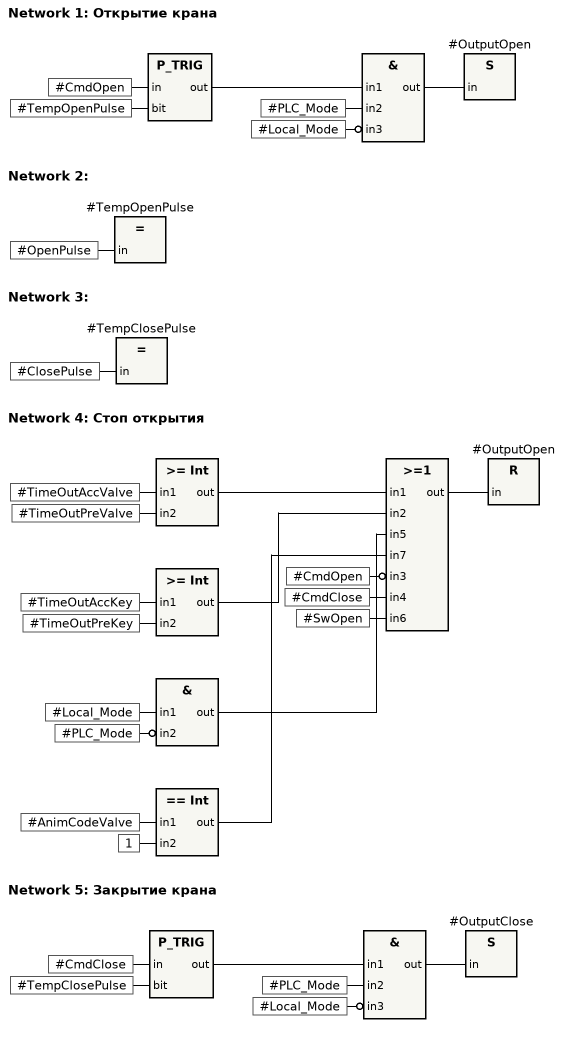
   #_w1 := #CmdOpen AND NOT #TempOpenPulse;   // rising edge
   #TempOpenPulse := #CmdOpen;
   IF #_w1 AND #PLC_Mode AND NOT #Local_Mode THEN #OutputOpen := TRUE; END_IF;
END_REGION

REGION Network 2
   #TempOpenPulse := #OpenPulse;
END_REGION

REGION Network 3
   #TempClosePulse := #ClosePulse;
END_REGION

REGION Network 4: Стоп открытия
   IF (#TimeOutAccValve >= #TimeOutPreValve) OR (#TimeOutAccKey >= #TimeOutPreKey) OR (#Local_Mode AND NOT #PLC_Mode) OR (#AnimCodeValve = 1) OR NOT #CmdOpen OR #CmdClose OR #SwOpen THEN
       #OutputOpen := FALSE;
   END_IF;
END_REGION

REGION Network 5: Закрытие крана
   #_w1 := #CmdClose AND NOT #TempClosePulse;   // rising edge
   #TempClosePulse := #CmdClose;
   IF #_w1 AND #PLC_Mode AND NOT #Local_Mode THEN #OutputClose := TRUE; END_IF;
END_REGION

REGION Network 6: Стоп закрытия
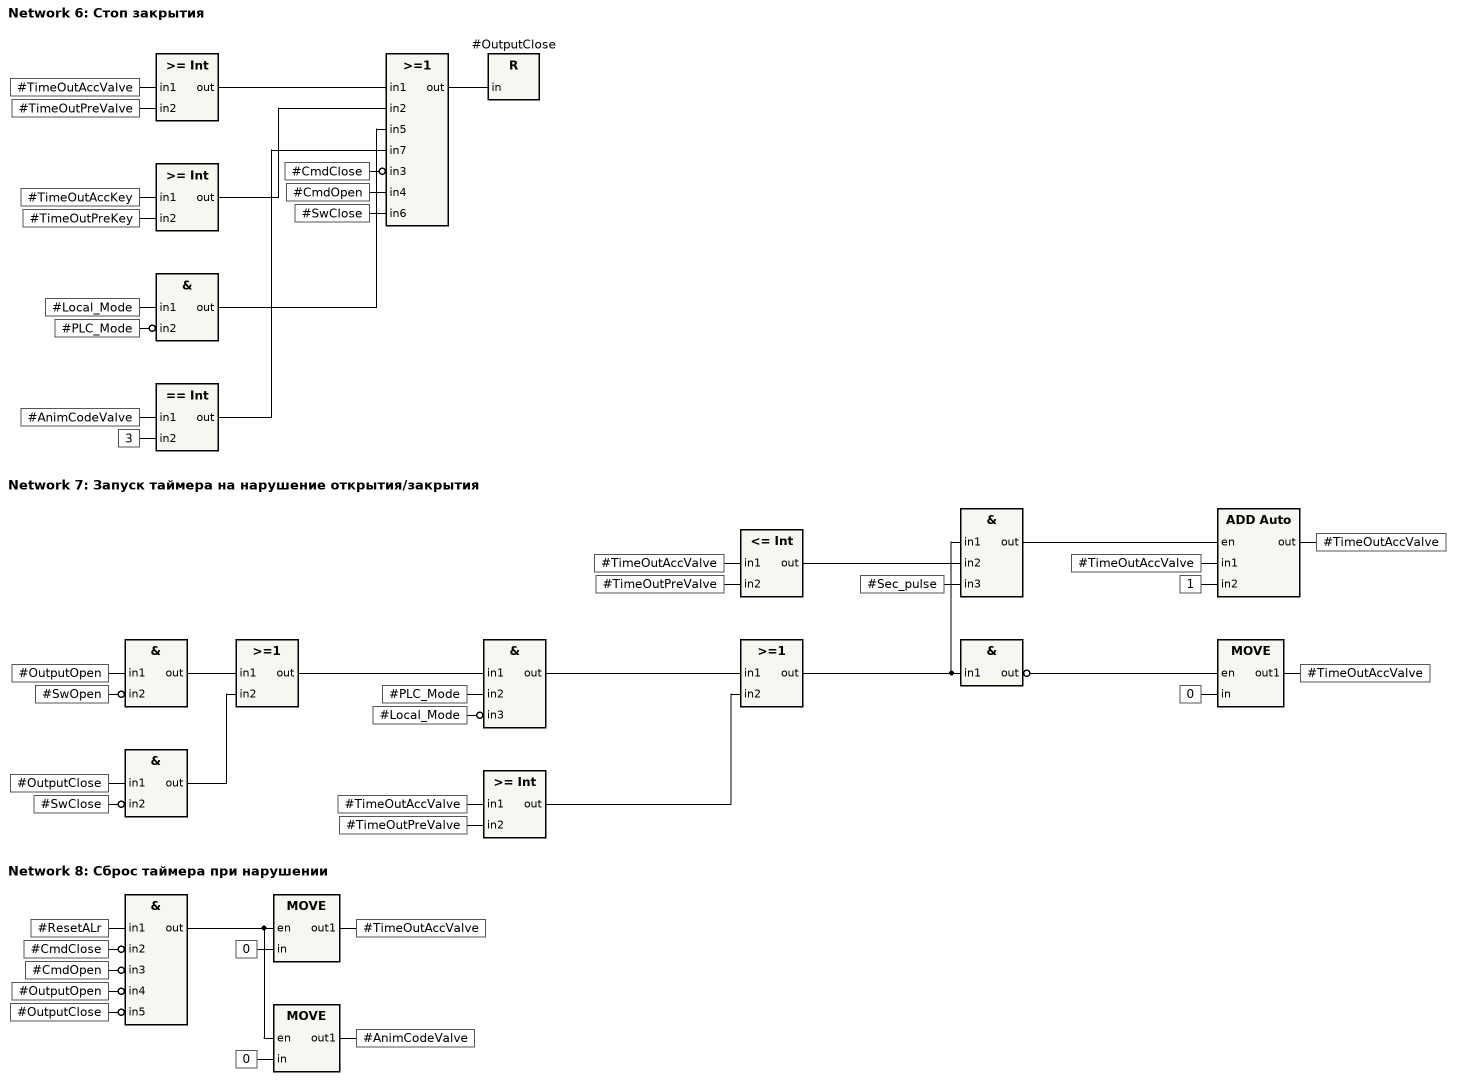
   IF (#TimeOutAccValve >= #TimeOutPreValve) OR (#TimeOutAccKey >= #TimeOutPreKey) OR (#Local_Mode AND NOT #PLC_Mode) OR (#AnimCodeValve = 3) OR NOT #CmdClose OR #CmdOpen OR #SwClose THEN
       #OutputClose := FALSE;
   END_IF;
END_REGION

REGION Network 7: Запуск таймера на нарушение открытия/закрытия
   #_w1 := (((#OutputOpen AND NOT #SwOpen) OR (#OutputClose AND NOT #SwClose)) AND #PLC_Mode AND NOT #Local_Mode) OR (#TimeOutAccValve >= #TimeOutPreValve);
   IF #_w1 AND (#TimeOutAccValve <= #TimeOutPreValve) AND #Sec_pulse THEN
       #TimeOutAccValve := #TimeOutAccValve + 1;
   END_IF;
   IF NOT #_w1 THEN #TimeOutAccValve := 0; END_IF;
END_REGION

REGION Network 8: Сброс таймера при нарушении
   IF #ResetALr AND NOT #CmdClose AND NOT #CmdOpen AND NOT #OutputOpen AND NOT #OutputClose THEN
       #TimeOutAccValve := 0;
       #AnimCodeValve := 0;
   END_IF;
END_REGION

REGION Network 9: Код анимации состояния крана
   // 0-Нейтральное
   // 1-Открыт
   // 2-Открывается
   // 3-Закрыт
   // 4-Закрывается
   // 10- Нарушения открытия
   // 11- Нарушения закрытия
   // 12- Открытие без команды
   // 13- Закрытие без команды
   // 14- Оба датчика включены
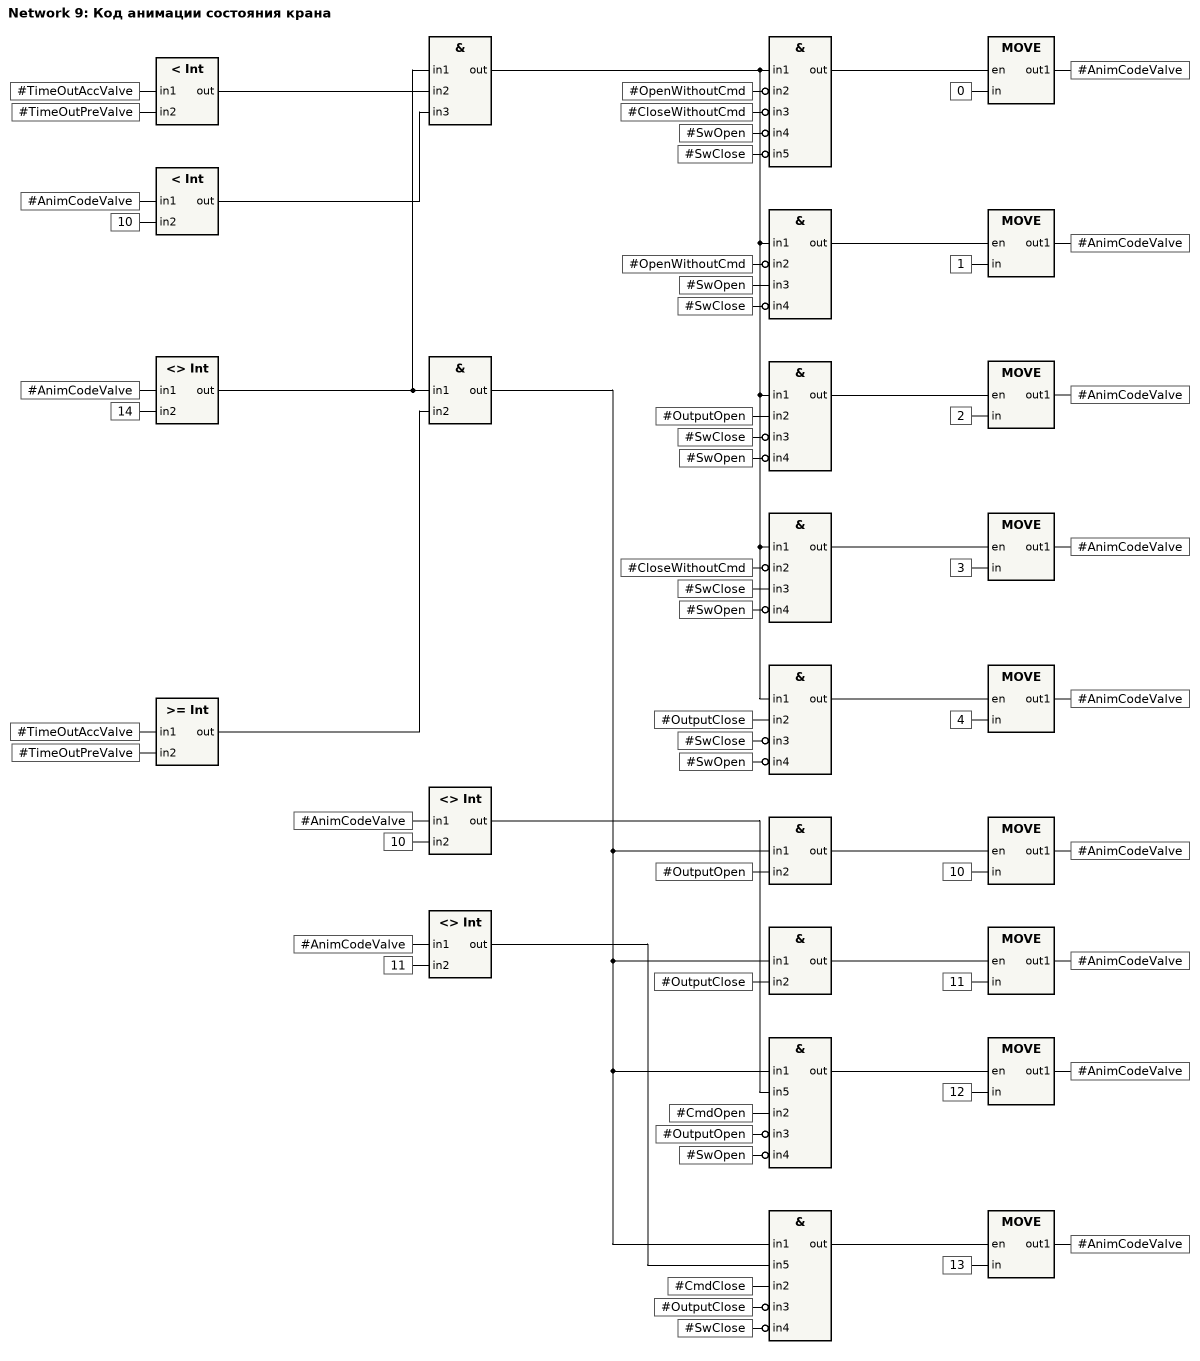
   #_w1 := #AnimCodeValve <> 14;
   #_w2 := #_w1 AND (#TimeOutAccValve < #TimeOutPreValve) AND (#AnimCodeValve < 10);
   IF #_w2 AND NOT #OpenWithoutCmd AND NOT #CloseWithoutCmd AND NOT #SwOpen AND NOT #SwClose THEN
       #AnimCodeValve := 0;
   END_IF;
   IF #_w2 AND NOT #OpenWithoutCmd AND #SwOpen AND NOT #SwClose THEN #AnimCodeValve := 1; END_IF;
   IF #_w2 AND #OutputOpen AND NOT #SwClose AND NOT #SwOpen THEN #AnimCodeValve := 2; END_IF;
   IF #_w2 AND NOT #CloseWithoutCmd AND #SwClose AND NOT #SwOpen THEN #AnimCodeValve := 3; END_IF;
   IF #_w2 AND #OutputClose AND NOT #SwClose AND NOT #SwOpen THEN #AnimCodeValve := 4; END_IF;
   #_w3 := #_w1 AND (#TimeOutAccValve >= #TimeOutPreValve);
   IF #_w3 AND #OutputOpen THEN #AnimCodeValve := 10; END_IF;
   IF #_w3 AND #OutputClose THEN #AnimCodeValve := 11; END_IF;
   IF #_w3 AND (#AnimCodeValve <> 10) AND #CmdOpen AND NOT #OutputOpen AND NOT #SwOpen THEN
       #AnimCodeValve := 12;
   END_IF;
   IF #_w3 AND (#AnimCodeValve <> 11) AND #CmdClose AND NOT #OutputClose AND NOT #SwClose THEN
       #AnimCodeValve := 13;
   END_IF;
END_REGION

REGION Network 10: Два датчика включены
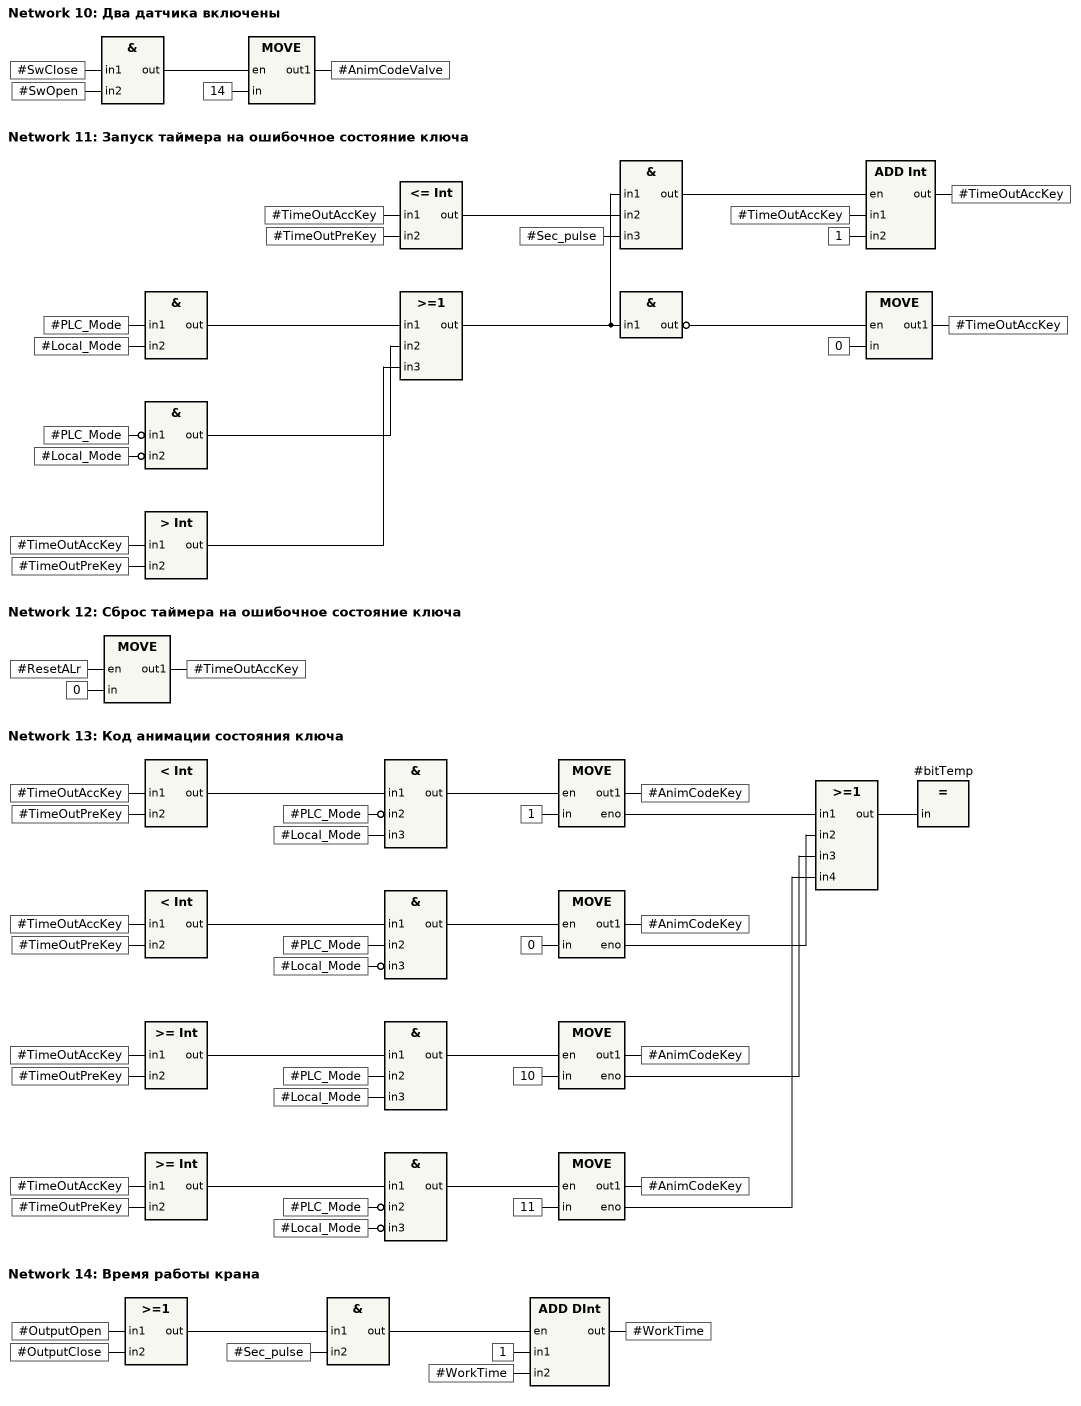
   IF #SwClose AND #SwOpen THEN #AnimCodeValve := 14; END_IF;
END_REGION

REGION Network 11: Запуск таймера на ошибочное состояние ключа
   #_w1 := (#PLC_Mode AND #Local_Mode) OR (NOT #PLC_Mode AND NOT #Local_Mode) OR (#TimeOutAccKey > #TimeOutPreKey);
   IF #_w1 AND (#TimeOutAccKey <= #TimeOutPreKey) AND #Sec_pulse THEN
       #TimeOutAccKey := #TimeOutAccKey + 1;
   END_IF;
   IF NOT #_w1 THEN #TimeOutAccKey := 0; END_IF;
END_REGION

REGION Network 12: Сброс таймера на ошибочное состояние ключа
   IF #ResetALr THEN #TimeOutAccKey := 0; END_IF;
END_REGION

REGION Network 13: Код анимации состояния ключа
   // ENO of a box is taken as its EN; it also drops when the box reports an error
   #_w1 := (#TimeOutAccKey < #TimeOutPreKey) AND NOT #PLC_Mode AND #Local_Mode;
   IF #_w1 THEN #AnimCodeKey := 1; END_IF;
   #_w2 := (#TimeOutAccKey < #TimeOutPreKey) AND #PLC_Mode AND NOT #Local_Mode;
   IF #_w2 THEN #AnimCodeKey := 0; END_IF;
   #_w3 := (#TimeOutAccKey >= #TimeOutPreKey) AND #PLC_Mode AND #Local_Mode;
   IF #_w3 THEN #AnimCodeKey := 10; END_IF;
   #_w4 := (#TimeOutAccKey >= #TimeOutPreKey) AND NOT #PLC_Mode AND NOT #Local_Mode;
   IF #_w4 THEN #AnimCodeKey := 11; END_IF;
   #bitTemp := #_w1 OR #_w2 OR #_w3 OR #_w4;
END_REGION

REGION Network 14: Время работы крана
   IF (#OutputOpen OR #OutputClose) AND #Sec_pulse THEN #WorkTime := 1 + #WorkTime; END_IF;
END_REGION

REGION Network 15: Сброс времени работы мотора
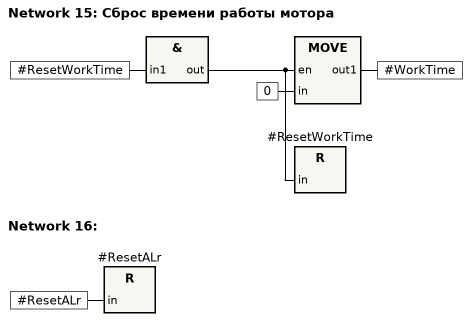
   IF #ResetWorkTime THEN
       #WorkTime := 0;
       #ResetWorkTime := FALSE;
   END_IF;
END_REGION

REGION Network 16
   IF #ResetALr THEN #ResetALr := FALSE; END_IF;
END_REGION
END_FUNCTION

FUNCTION "106_Analog_Type" : Void   // FC106, FBD
{ S7_Optimized_Access := 'TRUE' }
VERSION : 0.1
   VAR_INPUT
      Input : Int;
      Eng_Hi : Real;
      Eng_Lo : Real;
      Sp_HiHi : Real;
      Sp_Hi : Real;
      Sp_Lo : Real;
      Sp_LoLo : Real;
   END_VAR
   VAR_OUTPUT
      Value : Real;
      Alm_HiHi : Bool;
      Alm_Hi : Bool;
      Alm_Lo : Bool;
      Alm_LoLo : Bool;
      AnimCode : Int;
      OpenLoop : Bool;
      ShortCircuit : Bool;
   END_VAR
   VAR_TEMP
      Val_Conv : Real;
      Val_Temp : Real;
      Bool_Tmp : Bool;
      Input_Tmp : Int;
      tAlm_HiHi : Bool;
      tAlm_Hi : Bool;
      tAlm_Lo : Bool;
      tAlm_LoLo : Bool;
      tOpenLoop : Bool;
      tShortCircuit : Bool;
   END_VAR
BEGIN

REGION Network 1
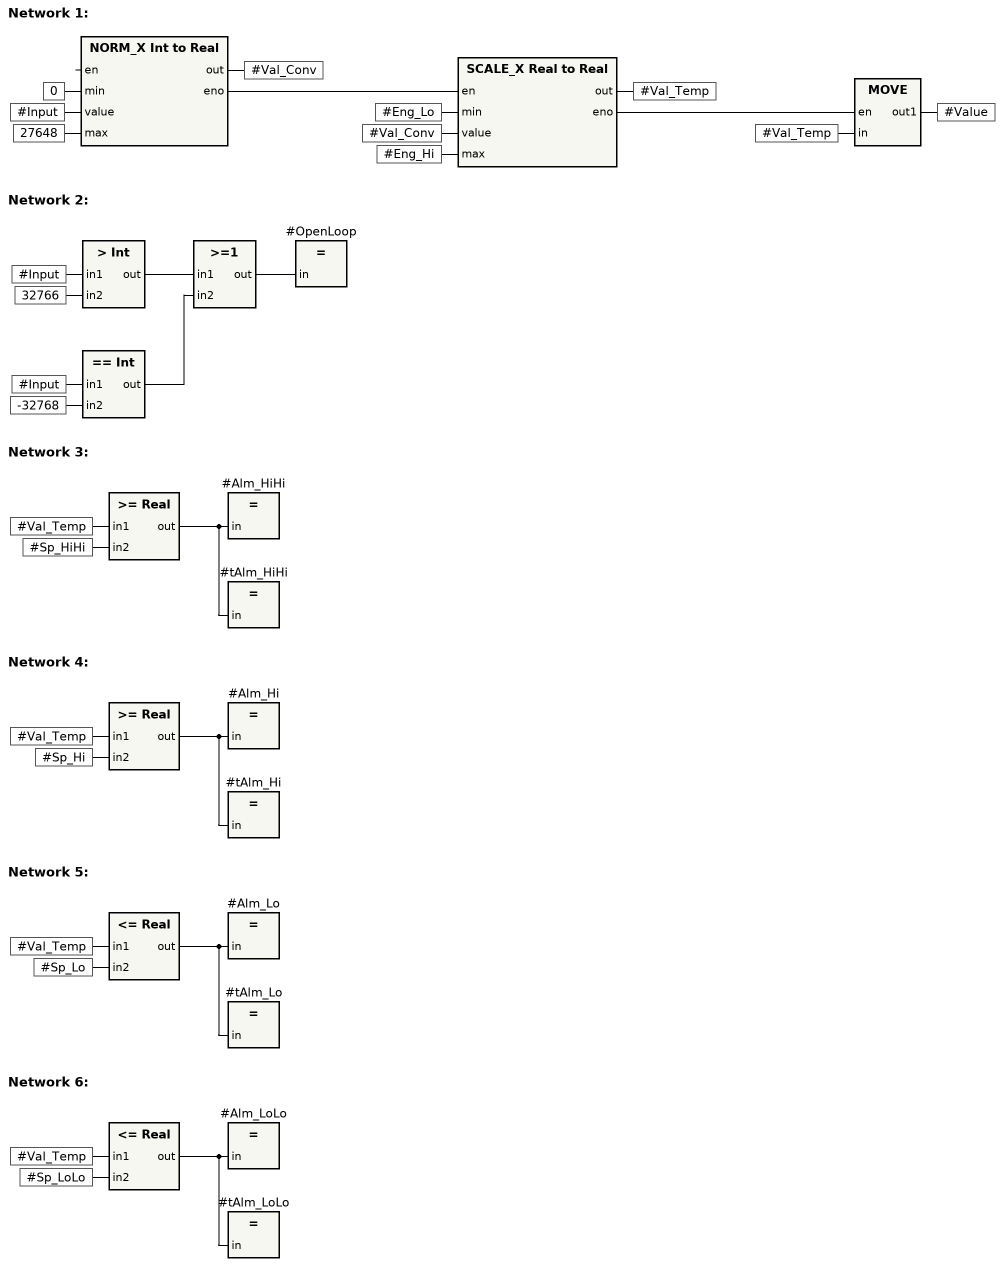
   // ENO of a box is taken as its EN; it also drops when the box reports an error
   #Val_Conv := NORM_X(MIN := 0, VALUE := #Input, MAX := 27648);
   #Val_Temp := SCALE_X(MIN := #Eng_Lo, VALUE := #Val_Conv, MAX := #Eng_Hi);
   #Value := #Val_Temp;
END_REGION

REGION Network 2
   #OpenLoop := (#Input > 32766) OR (#Input = (-32768));
END_REGION

REGION Network 3
   #Alm_HiHi := #Val_Temp >= #Sp_HiHi;
   #tAlm_HiHi := #Alm_HiHi;
END_REGION

REGION Network 4
   #Alm_Hi := #Val_Temp >= #Sp_Hi;
   #tAlm_Hi := #Alm_Hi;
END_REGION

REGION Network 5
   #Alm_Lo := #Val_Temp <= #Sp_Lo;
   #tAlm_Lo := #Alm_Lo;
END_REGION

REGION Network 6
   #Alm_LoLo := #Val_Temp <= #Sp_LoLo;
   #tAlm_LoLo := #Alm_LoLo;
END_REGION

REGION Network 7
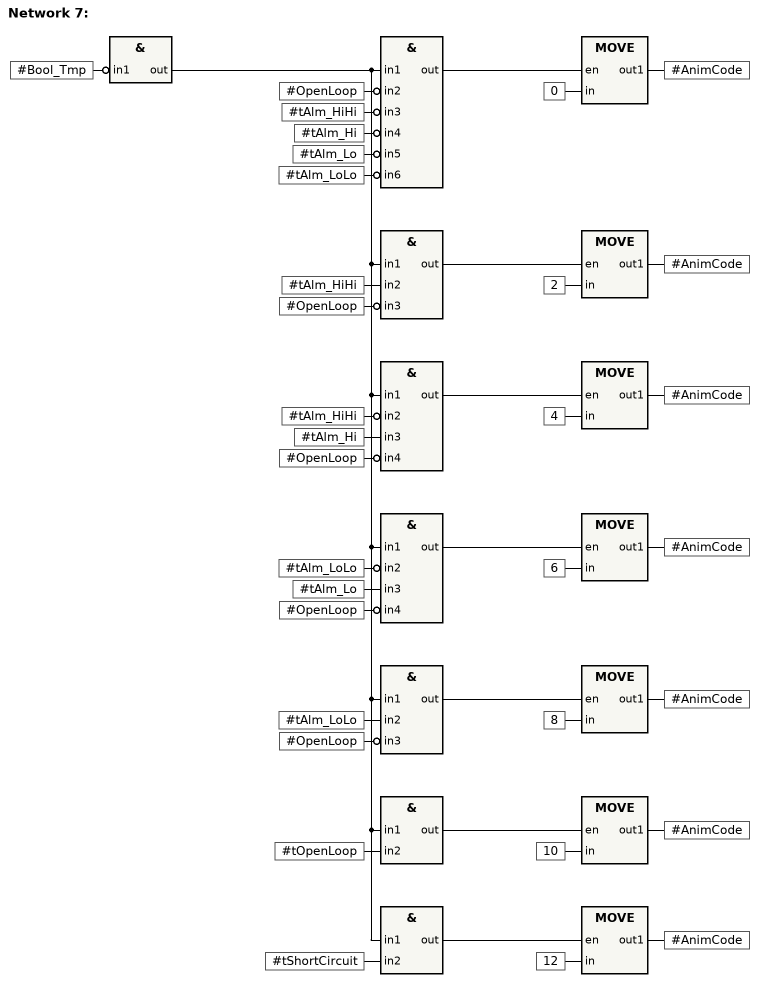
   IF NOT #Bool_Tmp AND NOT #OpenLoop AND NOT #tAlm_HiHi AND NOT #tAlm_Hi AND NOT #tAlm_Lo AND NOT #tAlm_LoLo THEN
       #AnimCode := 0;
   END_IF;
   IF NOT #Bool_Tmp AND #tAlm_HiHi AND NOT #OpenLoop THEN #AnimCode := 2; END_IF;
   IF NOT #Bool_Tmp AND NOT #tAlm_HiHi AND #tAlm_Hi AND NOT #OpenLoop THEN #AnimCode := 4; END_IF;
   IF NOT #Bool_Tmp AND NOT #tAlm_LoLo AND #tAlm_Lo AND NOT #OpenLoop THEN #AnimCode := 6; END_IF;
   IF NOT #Bool_Tmp AND #tAlm_LoLo AND NOT #OpenLoop THEN #AnimCode := 8; END_IF;
   IF NOT #Bool_Tmp AND #tOpenLoop THEN #AnimCode := 10; END_IF;
   IF NOT #Bool_Tmp AND #tShortCircuit THEN #AnimCode := 12; END_IF;
END_REGION
END_FUNCTION

ORGANIZATION_BLOCK "Main"   // OB1, LAD, ProgramCycle
TITLE = "Main Program Sweep (Cycle)"
{ S7_Optimized_Access := 'TRUE' }
VERSION : 0.1
   VAR_INPUT
      Initial_Call : Bool;   // Initial call of this OB
      Remanence : Bool;   // =True, if remanent data are available
   END_VAR
BEGIN

REGION Network 1
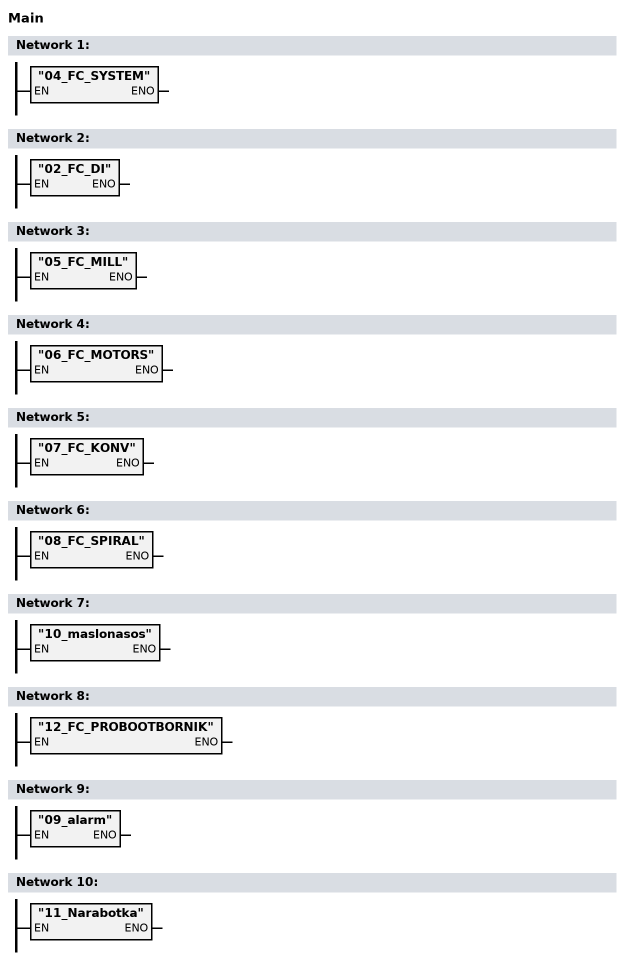
   RUNG wire#powerrail
      "04_FC_SYSTEM"()
   END_RUNG
   // the same network as SCL:
   "04_FC_SYSTEM"();
END_REGION

REGION Network 2
   RUNG wire#powerrail
      "02_FC_DI"()
   END_RUNG
   // the same network as SCL:
   "02_FC_DI"();
END_REGION

REGION Network 3
   RUNG wire#powerrail
      "05_FC_MILL"()
   END_RUNG
   // the same network as SCL:
   "05_FC_MILL"();
END_REGION

REGION Network 4
   RUNG wire#powerrail
      "06_FC_MOTORS"()
   END_RUNG
   // the same network as SCL:
   "06_FC_MOTORS"();
END_REGION

REGION Network 5
   RUNG wire#powerrail
      "07_FC_KONV"()
   END_RUNG
   // the same network as SCL:
   "07_FC_KONV"();
END_REGION

REGION Network 6
   RUNG wire#powerrail
      "08_FC_SPIRAL"()
   END_RUNG
   // the same network as SCL:
   "08_FC_SPIRAL"();
END_REGION

REGION Network 7
   RUNG wire#powerrail
      "10_maslonasos"()
   END_RUNG
   // the same network as SCL:
   "10_maslonasos"();
END_REGION

REGION Network 8
   RUNG wire#powerrail
      "12_FC_PROBOOTBORNIK"()
   END_RUNG
   // the same network as SCL:
   "12_FC_PROBOOTBORNIK"();
END_REGION

REGION Network 9
   RUNG wire#powerrail
      "09_alarm"()
   END_RUNG
   // the same network as SCL:
   "09_alarm"();
END_REGION

REGION Network 10
   RUNG wire#powerrail
      "11_Narabotka"()
   END_RUNG
   // the same network as SCL:
   "11_Narabotka"();
END_REGION
END_ORGANIZATION_BLOCK

ORGANIZATION_BLOCK "Time of day"   // OB10, LAD, TimeOfDay
{ S7_Optimized_Access := 'TRUE' }
VERSION : 0.1
   VAR_INPUT
      CaughtUp : Bool;   // OB call is caught up because time was set forward
      SecondTime : Bool;   // OB call is started a second time because time was set backward
   END_VAR
BEGIN
END_ORGANIZATION_BLOCK

ORGANIZATION_BLOCK "Time of day_1"   // OB11, LAD, TimeOfDay
{ S7_Optimized_Access := 'TRUE' }
VERSION : 0.1
   VAR_INPUT
      CaughtUp : Bool;   // OB call is caught up because time was set forward
      SecondTime : Bool;   // OB call is started a second time because time was set backward
   END_VAR
BEGIN
END_ORGANIZATION_BLOCK

ORGANIZATION_BLOCK "Cyclic interrupt"   // OB30, LAD, CyclicInterrupt
{ S7_Optimized_Access := 'TRUE' }
VERSION : 0.1
   VAR_INPUT
      Initial_Call : Bool;   // Initial call of this OB
      Event_Count : Int;   // Events discarded
   END_VAR
BEGIN

REGION Network 1
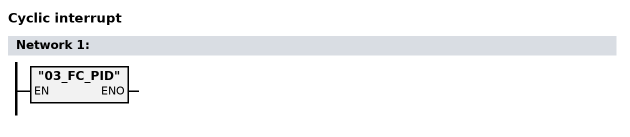
   RUNG wire#powerrail
      "03_FC_PID"()
   END_RUNG
   // the same network as SCL:
   "03_FC_PID"();
END_REGION
END_ORGANIZATION_BLOCK

ORGANIZATION_BLOCK "Cyclic interrupt_1"   // OB31, LAD, CyclicInterrupt
{ S7_Optimized_Access := 'TRUE' }
VERSION : 0.1
   VAR_INPUT
      Initial_Call : Bool;   // Initial call of this OB
      Event_Count : Int;   // Events discarded
   END_VAR
BEGIN

REGION Network 1
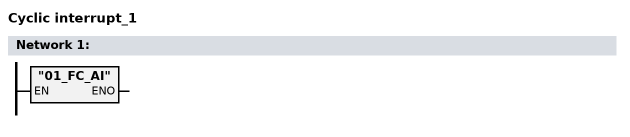
   RUNG wire#powerrail
      "01_FC_AI"()
   END_RUNG
   // the same network as SCL:
   "01_FC_AI"();
END_REGION
END_ORGANIZATION_BLOCK

ORGANIZATION_BLOCK "Cyclic interrupt_2"   // OB32, LAD, CyclicInterrupt
{ S7_Optimized_Access := 'TRUE' }
VERSION : 0.1
   VAR_INPUT
      Initial_Call : Bool;   // Initial call of this OB
      Event_Count : Int;   // Events discarded
   END_VAR
   VAR_TEMP
      r3s_tec : Real;
   END_VAR
BEGIN

REGION Network 1
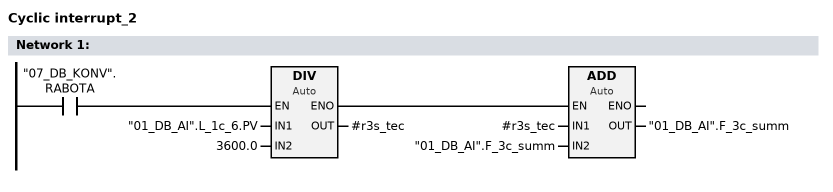
   RUNG wire#powerrail
      Contact( "07_DB_KONV".RABOTA )
      Div(in1 := "01_DB_AI".L_1c_6.PV, in2 := 3600.0, out => #r3s_tec)
      Add(in1 := #r3s_tec, in2 := "01_DB_AI".F_3c_summ, out => "01_DB_AI".F_3c_summ)
   END_RUNG
   // the same network as SCL:
   IF "07_DB_KONV".RABOTA THEN
       #r3s_tec := "01_DB_AI".L_1c_6.PV / 3600.0;
       "01_DB_AI".F_3c_summ := #r3s_tec + "01_DB_AI".F_3c_summ;
   END_IF;
END_REGION
END_ORGANIZATION_BLOCK

ORGANIZATION_BLOCK "Hardware interrupt"   // OB40, LAD, HWProcessInterrupt
{ S7_Optimized_Access := 'TRUE' }
VERSION : 0.1
   VAR_INPUT
      LADDR : Hw_Io;   // Hardware identifier
      USI : Word;   // User structure identifier
      IChannel : USInt;   // Interrupt channel number
      EventType : Byte;   // EventType
   END_VAR
BEGIN
END_ORGANIZATION_BLOCK

ORGANIZATION_BLOCK "Time error interrupt"   // OB80, LAD, TimeErrorInterrupt
{ S7_Optimized_Access := 'TRUE' }
VERSION : 0.1
   VAR_INPUT
      Fault_ID : Byte;   // Fault identifier
      Csg_OBnr : OB_Any;   // Number of OB causing the error
      Csg_Prio : UInt;   // Priority of OB causing the error
   END_VAR
BEGIN
END_ORGANIZATION_BLOCK

ORGANIZATION_BLOCK "Startup"   // OB100, LAD, Startup
TITLE = "Complete Restart"
{ S7_Optimized_Access := 'TRUE' }
VERSION : 0.1
   VAR_INPUT
      LostRetentive : Bool;   // True if retentive data are lost
      LostRTC : Bool;   // True if date and time are lost
   END_VAR
BEGIN
END_ORGANIZATION_BLOCK

ORGANIZATION_BLOCK "Main_1"   // OB123, LAD, ProgramCycle
TITLE = "Main Program Sweep (Cycle)"
{ S7_Optimized_Access := 'TRUE' }
VERSION : 0.1
   VAR_INPUT
      Initial_Call : Bool;   // Initial call of this OB
      Remanence : Bool;   // =True, if remanent data are available
   END_VAR
BEGIN
END_ORGANIZATION_BLOCK

(* ===== HMI "HMI_RT_1" =====
system functions are stored by id; their names below are inferred from use
connection "HMI_Соединение_1": ETHERNET, SMART_S7_1200_OMS

text list "ModeKlapan": 0 'Руч'; 1 'Авт'

text list "motor_AnimCode": 0 'Готов'; 1 'отключение'; 2 'Работа'; 4 'запуск'; 16 'нарушение'; 32 'нарушение'

text list "alarm_text_konv": 15 'Нарушение пуска'; 16 'Нарушение останова'; 17 'Уровен телеги'; 18 'Тросс выключатель'; 19 'Ток двигатель конвеера'; 20 ''

screen "memoscren" 1280x800
   IOField "Поле ввода-вывода_15" at 55,72 size 323x69; FormatPattern s999.9; Unit %
      ProcessValue <- "PV"
      Appearance <- "AnimCode"
   TextField "Text field_33" at 54,12 size 329x54; Text 'L_34'
   TextField "Text field_1" at 125,136 size 165x54; Text 'L12'
   TextField "Text field_2" at 126,252 size 162x54; Text 'L12'
   TextField "Text field_3" at 120,367 size 176x54; Text 'L12'
   IOField "Поле ввода-вывода_4" at 54,423 size 323x68; FormatPattern s999.9; Unit %
      ProcessValue <- "PV"
      Appearance <- "AnimCode"
   IOField "Поле ввода-вывода_5" at 55,303 size 317x70; FormatPattern s999.9; Unit %
      ProcessValue <- "PV"
      Appearance <- "AnimCode"
   IOField "Поле ввода-вывода_6" at 53,188 size 320x69; FormatPattern s999.9; Unit %
      ProcessValue <- "PV"
      Appearance <- "AnimCode"
   TextField "Text field_13" at 480,134 size 303x58; Text 'L12'
   TextField "Text field_19" at 476,370 size 304x58; Text 'L12'
   TextField "Text field_20" at 475,252 size 312x58; Text 'L12'
   TextField "Text field_21" at 921,258 size 267x47; Text 'L12'
   TextField "Text field_24" at 903,370 size 332x45; Text 'L12'
   IOField "Поле ввода-вывода_1" at 469,72 size 325x69; FormatPattern s999.9; Unit A
      ProcessValue <- "PV"
      Appearance <- "AnimCode"
   IOField "Поле ввода-вывода_2" at 464,186 size 325x65; FormatPattern s999.9; Unit A
      ProcessValue <- "PV"
      Appearance <- "AnimCode"
   IOField "Поле ввода-вывода_9" at 464,302 size 325x65; FormatPattern s999.9; Unit A
      ProcessValue <- "PV"
      Appearance <- "AnimCode"
   IOField "Поле ввода-вывода_12" at 898,417 size 340x70; FormatPattern s999.9; Unit %
      ProcessValue <- "PV"
      Appearance <- "AnimCode"
   IOField "Поле ввода-вывода_11" at 465,421 size 320x65; FormatPattern s999.9; Unit A
      ProcessValue <- "PV"
      Appearance <- "AnimCode"
   IOField "Поле ввода-вывода_3" at 898,302 size 340x70; FormatPattern s999.9; Unit %
      ProcessValue <- "PV"
      Appearance <- "AnimCode"
   TextField "Text field_5" at 467,11 size 332x58; Text 'L_34'
   TextField "Text field_29" at 1138,772 size 134x27; Text 'AI_param'
   TextField "Text field_9" at 889,773 size 134x27; Text 'Наработки'
   GraphicView "Graphic view_1" at 31,771 size 81x24; Picture "Left_Arrow"
   IOField "Поле ввода-вывода_7" at 903,71 size 323x64; FormatPattern s999.9; Unit %
      ProcessValue <- "PV"
      Appearance <- "AnimCode"
   TextField "Text field_11" at 845,16 size 415x54; Text 'L_34'
   IOField "Поле ввода-вывода_8" at 900,187 size 329x65; FormatPattern s999.9; Unit %
      ProcessValue <- "PV"
      Appearance <- "AnimCode"
   TextField "Text field_12" at 861,135 size 396x54; Text 'L12'
   Softkey "Softkey_F1" at 0,0 size 0x0
      on KeyDown: function_efd93a16()
   Softkey "Softkey_F10" at 0,0 size 0x0
      on KeyDown: ActivateScreen("ScreenParametr1", 0)
   Softkey "Softkey_F8" at 0,0 size 0x0
      on KeyDown: ActivateScreen("Naraboki", 0)